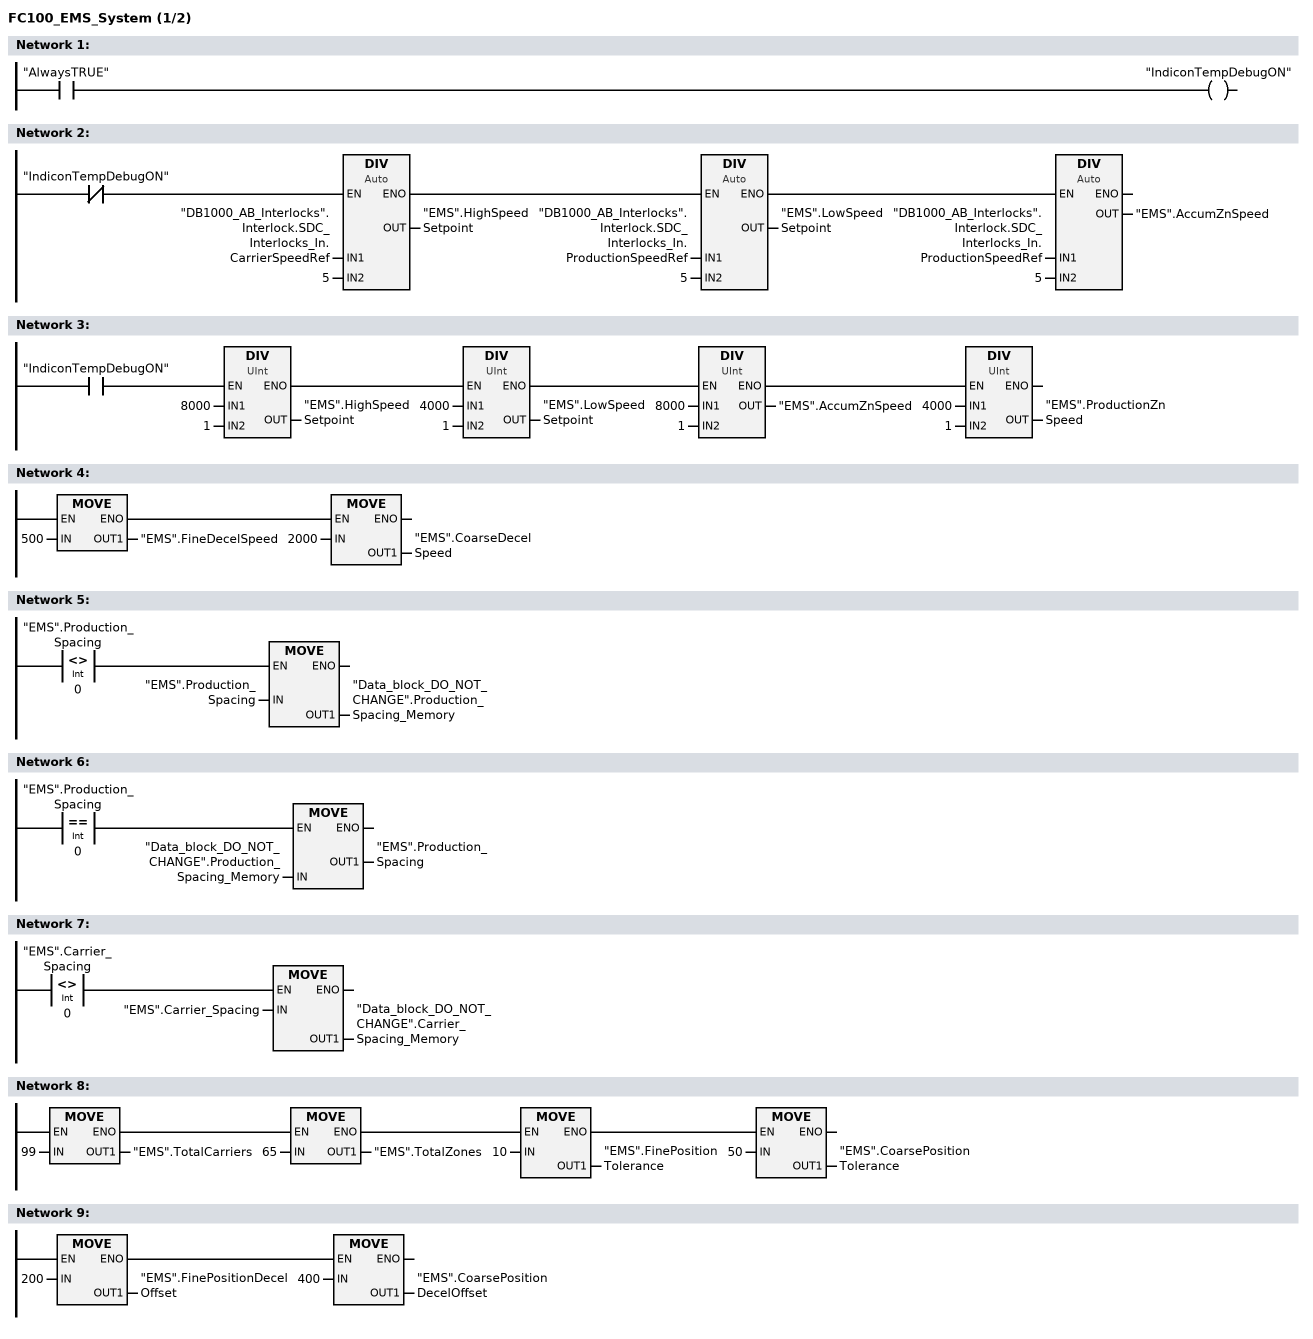
   RUNG wire#powerrail
      Contact( "AlwaysTRUE" )
      Coil( "IndiconTempDebugON" )
   END_RUNG
   // the same network as SCL:
   "IndiconTempDebugON" := "AlwaysTRUE";
END_REGION

REGION Network 2
   RUNG wire#powerrail
      I_Contact( "IndiconTempDebugON" )
      Div(in1 := "DB1000_AB_Interlocks".Interlock.SDC_Interlocks_In.CarrierSpeedRef, in2 := 5, out => "EMS".HighSpeedSetpoint)
      Div(in1 := "DB1000_AB_Interlocks".Interlock.SDC_Interlocks_In.ProductionSpeedRef, in2 := 5, out => "EMS".LowSpeedSetpoint)
      Div(in1 := "DB1000_AB_Interlocks".Interlock.SDC_Interlocks_In.ProductionSpeedRef, in2 := 5, out => "EMS".AccumZnSpeed)
   END_RUNG
   // the same network as SCL:
   IF NOT "IndiconTempDebugON" THEN
       "EMS".HighSpeedSetpoint := "DB1000_AB_Interlocks".Interlock.SDC_Interlocks_In.CarrierSpeedRef / 5;
       "EMS".LowSpeedSetpoint := "DB1000_AB_Interlocks".Interlock.SDC_Interlocks_In.ProductionSpeedRef / 5;
       "EMS".AccumZnSpeed := "DB1000_AB_Interlocks".Interlock.SDC_Interlocks_In.ProductionSpeedRef / 5;
   END_IF;
END_REGION

REGION Network 3
   RUNG wire#powerrail
      Contact( "IndiconTempDebugON" )
      { S7_Templates := "SrcType := UInt" } Div(in1 := 8000, in2 := 1, out => "EMS".HighSpeedSetpoint)
      { S7_Templates := "SrcType := UInt" } Div(in1 := 4000, in2 := 1, out => "EMS".LowSpeedSetpoint)
      { S7_Templates := "SrcType := UInt" } Div(in1 := 8000, in2 := 1, out => "EMS".AccumZnSpeed)
      { S7_Templates := "SrcType := UInt" } Div(in1 := 4000, in2 := 1, out => "EMS".ProductionZnSpeed)
   END_RUNG
   // the same network as SCL:
   IF "IndiconTempDebugON" THEN
       "EMS".HighSpeedSetpoint := 8000 / 1;
       "EMS".LowSpeedSetpoint := 4000 / 1;
       "EMS".AccumZnSpeed := 8000 / 1;
       "EMS".ProductionZnSpeed := 4000 / 1;
   END_IF;
END_REGION

REGION Network 4
   RUNG wire#powerrail
      Move(in := 500, out1 => "EMS".FineDecelSpeed)
      Move(in := 2000, out1 => "EMS".CoarseDecelSpeed)
   END_RUNG
   // the same network as SCL:
   "EMS".FineDecelSpeed := 500;
   "EMS".CoarseDecelSpeed := 2000;
END_REGION

REGION Network 5
   RUNG wire#powerrail
      { S7_Templates := "SrcType := Int" } NE_Contact(in1 := "EMS".Production_Spacing, in2 := 0)
      Move(in := "EMS".Production_Spacing, out1 => "Data_block_DO_NOT_CHANGE".Production_Spacing_Memory)
   END_RUNG
   // the same network as SCL:
   IF "EMS".Production_Spacing <> 0 THEN
       "Data_block_DO_NOT_CHANGE".Production_Spacing_Memory := "EMS".Production_Spacing;
   END_IF;
END_REGION

REGION Network 6
   RUNG wire#powerrail
      { S7_Templates := "SrcType := Int" } EQ_Contact(in1 := "EMS".Production_Spacing, in2 := 0)
      Move(in := "Data_block_DO_NOT_CHANGE".Production_Spacing_Memory, out1 => "EMS".Production_Spacing)
   END_RUNG
   // the same network as SCL:
   IF "EMS".Production_Spacing = 0 THEN
       "EMS".Production_Spacing := "Data_block_DO_NOT_CHANGE".Production_Spacing_Memory;
   END_IF;
END_REGION

REGION Network 7
   RUNG wire#powerrail
      { S7_Templates := "SrcType := Int" } NE_Contact(in1 := "EMS".Carrier_Spacing, in2 := 0)
      Move(in := "EMS".Carrier_Spacing, out1 => "Data_block_DO_NOT_CHANGE".Carrier_Spacing_Memory)
   END_RUNG
   // the same network as SCL:
   IF "EMS".Carrier_Spacing <> 0 THEN
       "Data_block_DO_NOT_CHANGE".Carrier_Spacing_Memory := "EMS".Carrier_Spacing;
   END_IF;
END_REGION

REGION Network 8
   RUNG wire#powerrail
      Move(in := 99, out1 => "EMS".TotalCarriers)
      Move(in := 65, out1 => "EMS".TotalZones)
      Move(in := 10, out1 => "EMS".FinePositionTolerance)
      Move(in := 50, out1 => "EMS".CoarsePositionTolerance)
   END_RUNG
   // the same network as SCL:
   "EMS".TotalCarriers := 99;
   "EMS".TotalZones := 65;
   "EMS".FinePositionTolerance := 10;
   "EMS".CoarsePositionTolerance := 50;
END_REGION

REGION Network 9
   RUNG wire#powerrail
      Move(in := 200, out1 => "EMS".FinePositionDecelOffset)
      Move(in := 400, out1 => "EMS".CoarsePositionDecelOffset)
   END_RUNG
   // the same network as SCL:
   "EMS".FinePositionDecelOffset := 200;
   "EMS".CoarsePositionDecelOffset := 400;
END_REGION

REGION Network 10
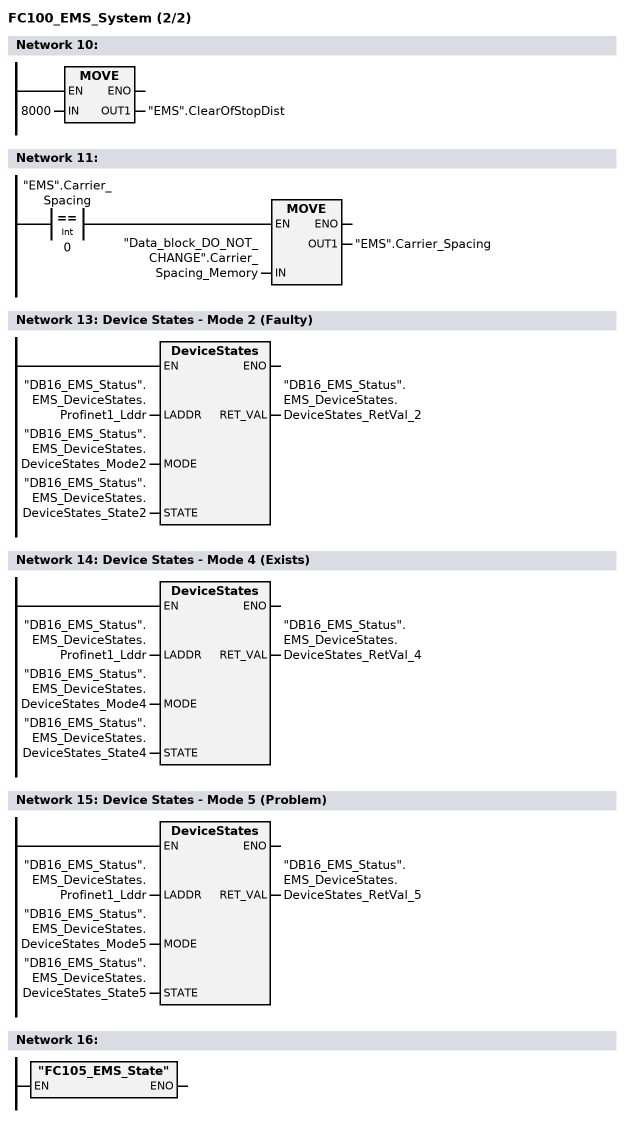
   RUNG wire#powerrail
      Move(in := 8000, out1 => "EMS".ClearOfStopDist)
   END_RUNG
   // the same network as SCL:
   "EMS".ClearOfStopDist := 8000;
END_REGION

REGION Network 11
   RUNG wire#powerrail
      { S7_Templates := "SrcType := Int" } EQ_Contact(in1 := "EMS".Carrier_Spacing, in2 := 0)
      Move(in := "Data_block_DO_NOT_CHANGE".Carrier_Spacing_Memory, out1 => "EMS".Carrier_Spacing)
   END_RUNG
   // the same network as SCL:
   IF "EMS".Carrier_Spacing = 0 THEN
       "EMS".Carrier_Spacing := "Data_block_DO_NOT_CHANGE".Carrier_Spacing_Memory;
   END_IF;
END_REGION

REGION Network 13: Device States - Mode 2 (Faulty)
   // no SCL statement known for DeviceStates: written as a call
   "DB16_EMS_Status".EMS_DeviceStates.DeviceStates_RetVal_2 := DeviceStates(LADDR := "DB16_EMS_Status".EMS_DeviceStates.Profinet1_Lddr,
                           MODE := "DB16_EMS_Status".EMS_DeviceStates.DeviceStates_Mode2,
                           STATE := "DB16_EMS_Status".EMS_DeviceStates.DeviceStates_State2);
END_REGION

REGION Network 14: Device States - Mode 4 (Exists)
   // no SCL statement known for DeviceStates: written as a call
   "DB16_EMS_Status".EMS_DeviceStates.DeviceStates_RetVal_4 := DeviceStates(LADDR := "DB16_EMS_Status".EMS_DeviceStates.Profinet1_Lddr,
                           MODE := "DB16_EMS_Status".EMS_DeviceStates.DeviceStates_Mode4,
                           STATE := "DB16_EMS_Status".EMS_DeviceStates.DeviceStates_State4);
END_REGION

REGION Network 15: Device States - Mode 5 (Problem)
   // no SCL statement known for DeviceStates: written as a call
   "DB16_EMS_Status".EMS_DeviceStates.DeviceStates_RetVal_5 := DeviceStates(LADDR := "DB16_EMS_Status".EMS_DeviceStates.Profinet1_Lddr,
                           MODE := "DB16_EMS_Status".EMS_DeviceStates.DeviceStates_Mode5,
                           STATE := "DB16_EMS_Status".EMS_DeviceStates.DeviceStates_State5);
END_REGION

REGION Network 16
   RUNG wire#powerrail
      "FC105_EMS_State"()
   END_RUNG
   // the same network as SCL:
   "FC105_EMS_State"();
END_REGION
END_FUNCTION

FUNCTION "FC102_TCop_Map_SDCOut" : Void   // FC102, LAD
{ S7_Optimized_Access := 'TRUE' }
VERSION : 0.1
   VAR_TEMP
      tempdisplay : Bool;
      TotalCarriers : Int;
      TotalZones : Int;
      OneShot : Bool;
      countpulse : Bool;
   END_VAR
   VAR_TEMP   // added for the SCL form of the ladder/FBD networks
      _w1 : Bool;
   END_VAR
BEGIN

REGION Network 1
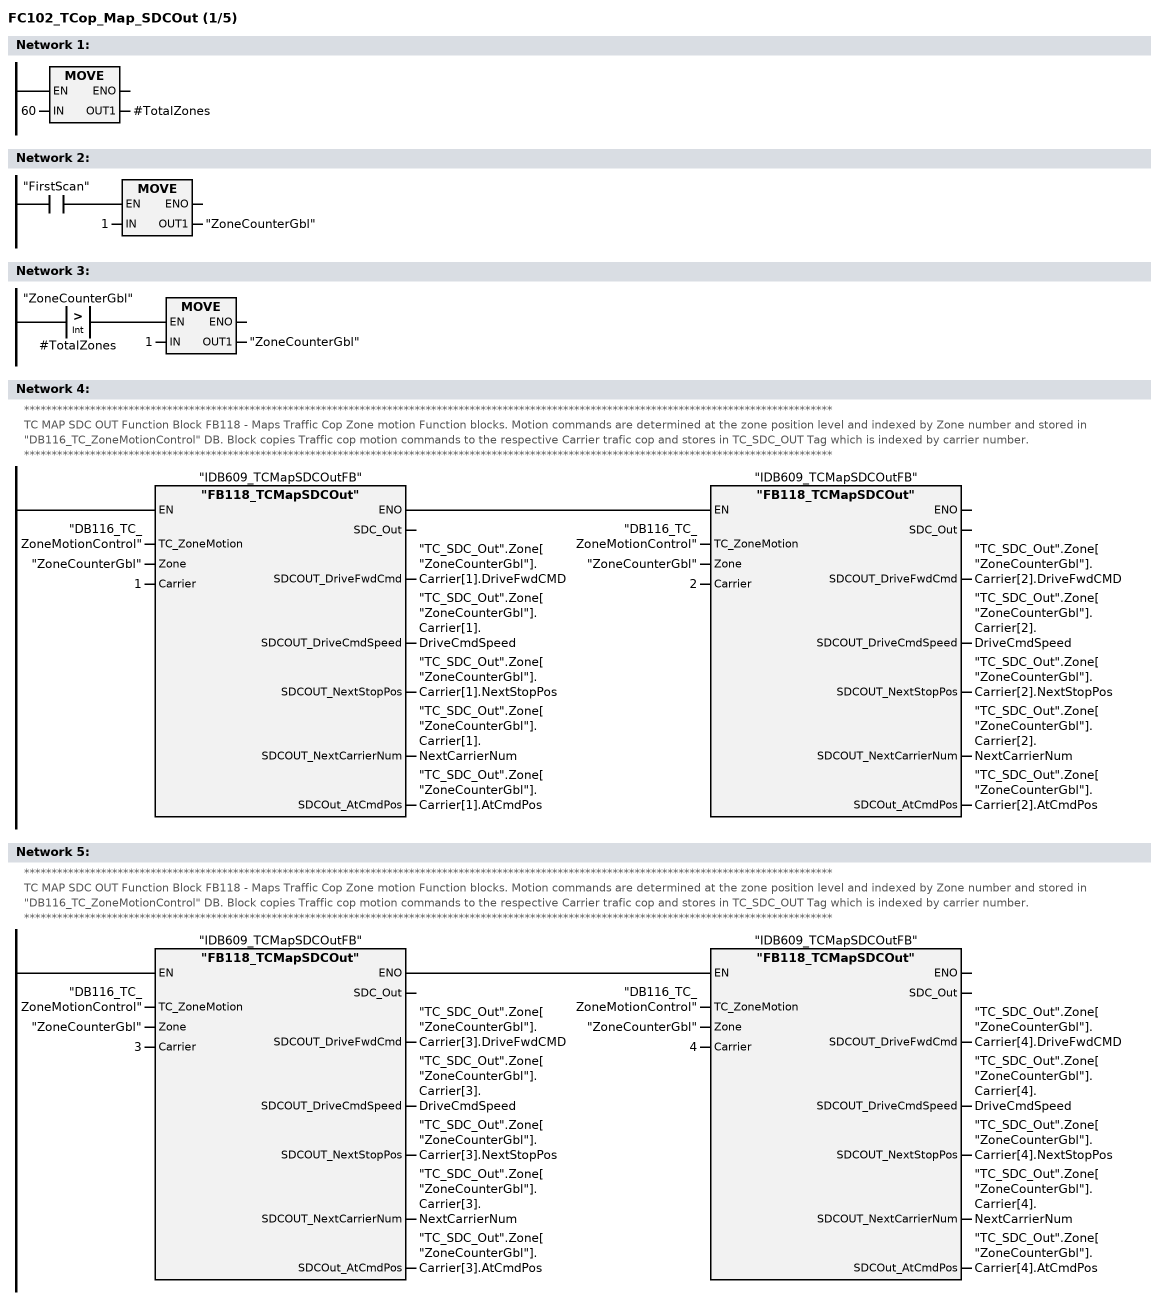
   RUNG wire#powerrail
      Move(in := 60, out1 => #TotalZones)
   END_RUNG
   // the same network as SCL:
   #TotalZones := 60;
END_REGION

REGION Network 2
   RUNG wire#powerrail
      Contact( "FirstScan" )
      Move(in := 1, out1 => "ZoneCounterGbl")
   END_RUNG
   // the same network as SCL:
   IF "FirstScan" THEN "ZoneCounterGbl" := 1; END_IF;
END_REGION

REGION Network 3
   RUNG wire#powerrail
      { S7_Templates := "SrcType := Int" } GT_Contact(in1 := "ZoneCounterGbl", in2 := #TotalZones)
      Move(in := 1, out1 => "ZoneCounterGbl")
   END_RUNG
   // the same network as SCL:
   IF "ZoneCounterGbl" > #TotalZones THEN "ZoneCounterGbl" := 1; END_IF;
END_REGION

REGION Network 4
   // ***************************************************************************************************************************************************
   // 
   // TC MAP SDC OUT Function Block FB118 - Maps Traffic Cop Zone motion Function blocks. Motion commands are determined at the zone position level and indexed by Zone number and stored in 
   //  "DB116_TC_ZoneMotionControl" DB. Block copies Traffic cop motion commands to the respective Carrier trafic cop and stores in TC_SDC_OUT Tag which is indexed by carrier number. 
   // 
   // ***************************************************************************************************************************************************
   RUNG wire#powerrail
      "IDB609_TCMapSDCOutFB"(TC_ZoneMotion := "DB116_TC_ZoneMotionControl", Zone := "ZoneCounterGbl", Carrier := 1, SDC_Out =>, SDCOUT_DriveFwdCmd => "TC_SDC_Out".Zone["ZoneCounterGbl"].Carrier[1].DriveFwdCMD, SDCOUT_DriveCmdSpeed => "TC_SDC_Out".Zone["ZoneCounterGbl"].Carrier[1].DriveCmdSpeed, SDCOUT_NextStopPos => "TC_SDC_Out".Zone["ZoneCounterGbl"].Carrier[1].NextStopPos, SDCOUT_NextCarrierNum => "TC_SDC_Out".Zone["ZoneCounterGbl"].Carrier[1].NextCarrierNum, SDCOut_AtCmdPos => "TC_SDC_Out".Zone["ZoneCounterGbl"].Carrier[1].AtCmdPos)
      "IDB609_TCMapSDCOutFB"(TC_ZoneMotion := "DB116_TC_ZoneMotionControl", Zone := "ZoneCounterGbl", Carrier := 2, SDC_Out =>, SDCOUT_DriveFwdCmd => "TC_SDC_Out".Zone["ZoneCounterGbl"].Carrier[2].DriveFwdCMD, SDCOUT_DriveCmdSpeed => "TC_SDC_Out".Zone["ZoneCounterGbl"].Carrier[2].DriveCmdSpeed, SDCOUT_NextStopPos => "TC_SDC_Out".Zone["ZoneCounterGbl"].Carrier[2].NextStopPos, SDCOUT_NextCarrierNum => "TC_SDC_Out".Zone["ZoneCounterGbl"].Carrier[2].NextCarrierNum, SDCOut_AtCmdPos => "TC_SDC_Out".Zone["ZoneCounterGbl"].Carrier[2].AtCmdPos)
   END_RUNG
   // the same network as SCL:
   "IDB609_TCMapSDCOutFB"(TC_ZoneMotion := "DB116_TC_ZoneMotionControl",   // "FB118_TCMapSDCOut"
                          Zone := "ZoneCounterGbl",
                          Carrier := 1,
                          SDCOUT_DriveFwdCmd => "TC_SDC_Out".Zone["ZoneCounterGbl"].Carrier[1].DriveFwdCMD,
                          SDCOUT_DriveCmdSpeed => "TC_SDC_Out".Zone["ZoneCounterGbl"].Carrier[1].DriveCmdSpeed,
                          SDCOUT_NextStopPos => "TC_SDC_Out".Zone["ZoneCounterGbl"].Carrier[1].NextStopPos,
                          SDCOUT_NextCarrierNum => "TC_SDC_Out".Zone["ZoneCounterGbl"].Carrier[1].NextCarrierNum,
                          SDCOut_AtCmdPos => "TC_SDC_Out".Zone["ZoneCounterGbl"].Carrier[1].AtCmdPos,
                          ENO => #_w1);
   IF #_w1 THEN
       "IDB609_TCMapSDCOutFB"(TC_ZoneMotion := "DB116_TC_ZoneMotionControl",   // "FB118_TCMapSDCOut"
                              Zone := "ZoneCounterGbl",
                              Carrier := 2,
                              SDCOUT_DriveFwdCmd => "TC_SDC_Out".Zone["ZoneCounterGbl"].Carrier[2].DriveFwdCMD,
                              SDCOUT_DriveCmdSpeed => "TC_SDC_Out".Zone["ZoneCounterGbl"].Carrier[2].DriveCmdSpeed,
                              SDCOUT_NextStopPos => "TC_SDC_Out".Zone["ZoneCounterGbl"].Carrier[2].NextStopPos,
                              SDCOUT_NextCarrierNum => "TC_SDC_Out".Zone["ZoneCounterGbl"].Carrier[2].NextCarrierNum,
                              SDCOut_AtCmdPos => "TC_SDC_Out".Zone["ZoneCounterGbl"].Carrier[2].AtCmdPos);
   END_IF;
END_REGION

REGION Network 5
   // ***************************************************************************************************************************************************
   // 
   // TC MAP SDC OUT Function Block FB118 - Maps Traffic Cop Zone motion Function blocks. Motion commands are determined at the zone position level and indexed by Zone number and stored in 
   //  "DB116_TC_ZoneMotionControl" DB. Block copies Traffic cop motion commands to the respective Carrier trafic cop and stores in TC_SDC_OUT Tag which is indexed by carrier number. 
   // 
   // ***************************************************************************************************************************************************
   RUNG wire#powerrail
      "IDB609_TCMapSDCOutFB"(TC_ZoneMotion := "DB116_TC_ZoneMotionControl", Zone := "ZoneCounterGbl", Carrier := 3, SDC_Out =>, SDCOUT_DriveFwdCmd => "TC_SDC_Out".Zone["ZoneCounterGbl"].Carrier[3].DriveFwdCMD, SDCOUT_DriveCmdSpeed => "TC_SDC_Out".Zone["ZoneCounterGbl"].Carrier[3].DriveCmdSpeed, SDCOUT_NextStopPos => "TC_SDC_Out".Zone["ZoneCounterGbl"].Carrier[3].NextStopPos, SDCOUT_NextCarrierNum => "TC_SDC_Out".Zone["ZoneCounterGbl"].Carrier[3].NextCarrierNum, SDCOut_AtCmdPos => "TC_SDC_Out".Zone["ZoneCounterGbl"].Carrier[3].AtCmdPos)
      "IDB609_TCMapSDCOutFB"(TC_ZoneMotion := "DB116_TC_ZoneMotionControl", Zone := "ZoneCounterGbl", Carrier := 4, SDC_Out =>, SDCOUT_DriveFwdCmd => "TC_SDC_Out".Zone["ZoneCounterGbl"].Carrier[4].DriveFwdCMD, SDCOUT_DriveCmdSpeed => "TC_SDC_Out".Zone["ZoneCounterGbl"].Carrier[4].DriveCmdSpeed, SDCOUT_NextStopPos => "TC_SDC_Out".Zone["ZoneCounterGbl"].Carrier[4].NextStopPos, SDCOUT_NextCarrierNum => "TC_SDC_Out".Zone["ZoneCounterGbl"].Carrier[4].NextCarrierNum, SDCOut_AtCmdPos => "TC_SDC_Out".Zone["ZoneCounterGbl"].Carrier[4].AtCmdPos)
   END_RUNG
   // the same network as SCL:
   "IDB609_TCMapSDCOutFB"(TC_ZoneMotion := "DB116_TC_ZoneMotionControl",   // "FB118_TCMapSDCOut"
                          Zone := "ZoneCounterGbl",
                          Carrier := 3,
                          SDCOUT_DriveFwdCmd => "TC_SDC_Out".Zone["ZoneCounterGbl"].Carrier[3].DriveFwdCMD,
                          SDCOUT_DriveCmdSpeed => "TC_SDC_Out".Zone["ZoneCounterGbl"].Carrier[3].DriveCmdSpeed,
                          SDCOUT_NextStopPos => "TC_SDC_Out".Zone["ZoneCounterGbl"].Carrier[3].NextStopPos,
                          SDCOUT_NextCarrierNum => "TC_SDC_Out".Zone["ZoneCounterGbl"].Carrier[3].NextCarrierNum,
                          SDCOut_AtCmdPos => "TC_SDC_Out".Zone["ZoneCounterGbl"].Carrier[3].AtCmdPos,
                          ENO => #_w1);
   IF #_w1 THEN
       "IDB609_TCMapSDCOutFB"(TC_ZoneMotion := "DB116_TC_ZoneMotionControl",   // "FB118_TCMapSDCOut"
                              Zone := "ZoneCounterGbl",
                              Carrier := 4,
                              SDCOUT_DriveFwdCmd => "TC_SDC_Out".Zone["ZoneCounterGbl"].Carrier[4].DriveFwdCMD,
                              SDCOUT_DriveCmdSpeed => "TC_SDC_Out".Zone["ZoneCounterGbl"].Carrier[4].DriveCmdSpeed,
                              SDCOUT_NextStopPos => "TC_SDC_Out".Zone["ZoneCounterGbl"].Carrier[4].NextStopPos,
                              SDCOUT_NextCarrierNum => "TC_SDC_Out".Zone["ZoneCounterGbl"].Carrier[4].NextCarrierNum,
                              SDCOut_AtCmdPos => "TC_SDC_Out".Zone["ZoneCounterGbl"].Carrier[4].AtCmdPos);
   END_IF;
END_REGION

REGION Network 6
   // ***************************************************************************************************************************************************
   // 
   // TC MAP SDC OUT Function Block FB118 - Maps Traffic Cop Zone motion Function blocks. Motion commands are determined at the zone position level and indexed by Zone number and stored in 
   //  "DB116_TC_ZoneMotionControl" DB. Block copies Traffic cop motion commands to the respective Carrier trafic cop and stores in TC_SDC_OUT Tag which is indexed by carrier number. 
   // 
   // ***************************************************************************************************************************************************
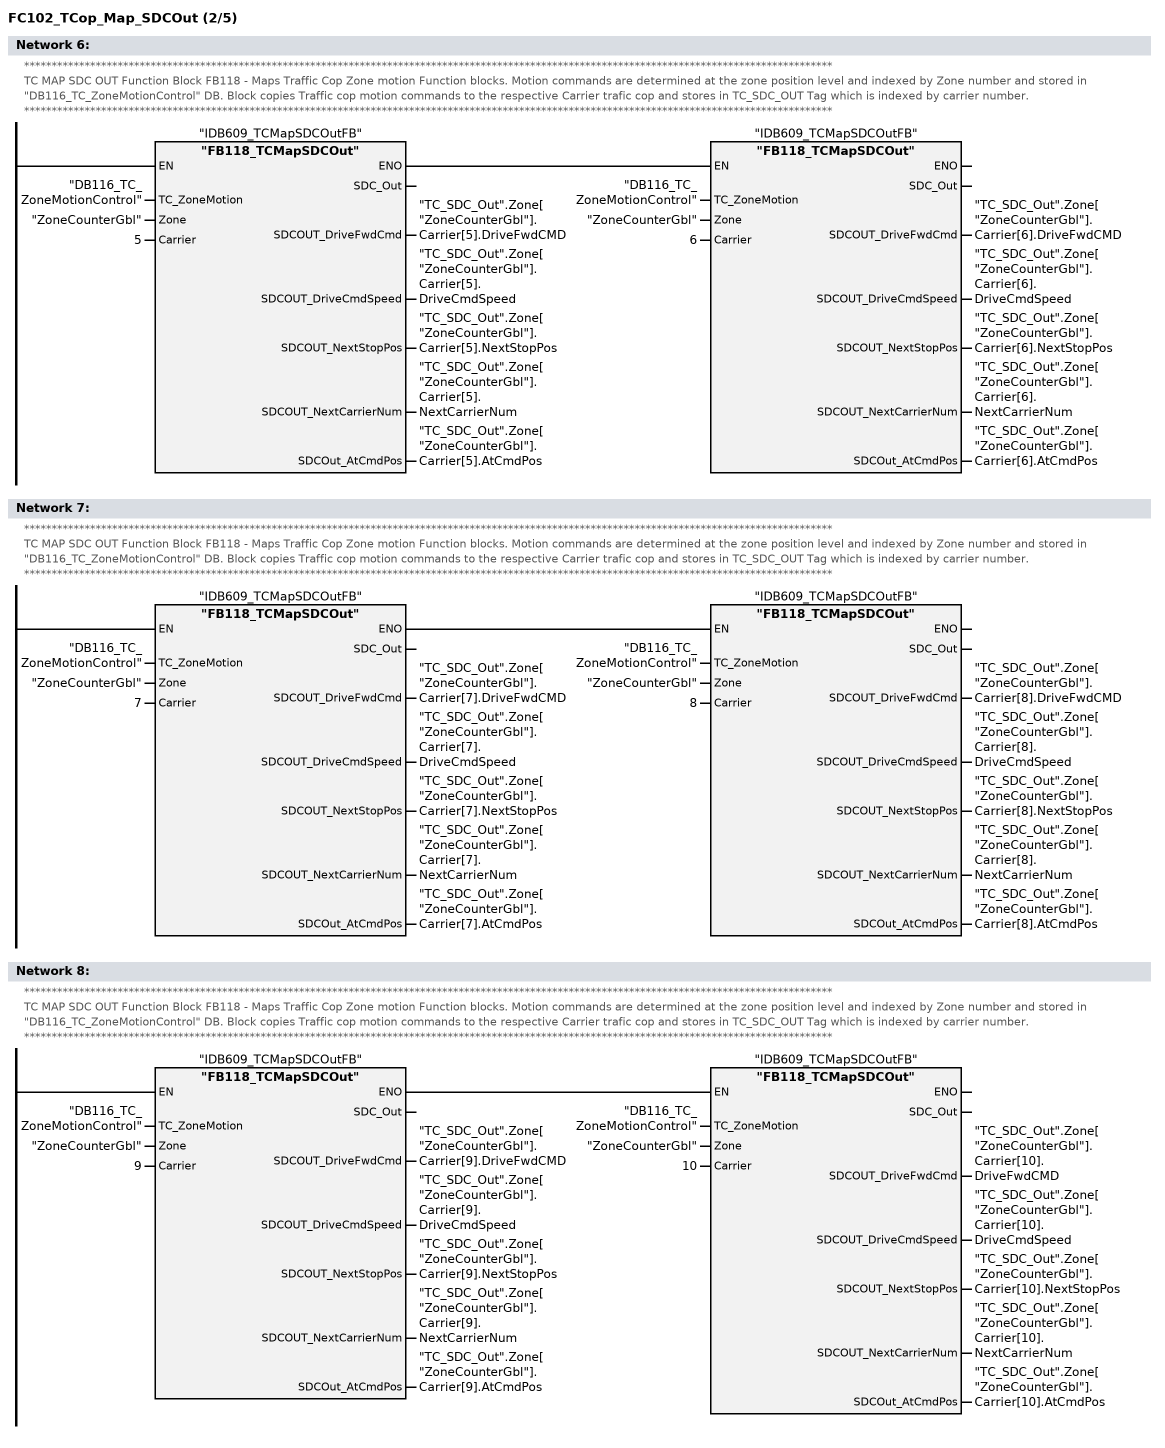
   RUNG wire#powerrail
      "IDB609_TCMapSDCOutFB"(TC_ZoneMotion := "DB116_TC_ZoneMotionControl", Zone := "ZoneCounterGbl", Carrier := 5, SDC_Out =>, SDCOUT_DriveFwdCmd => "TC_SDC_Out".Zone["ZoneCounterGbl"].Carrier[5].DriveFwdCMD, SDCOUT_DriveCmdSpeed => "TC_SDC_Out".Zone["ZoneCounterGbl"].Carrier[5].DriveCmdSpeed, SDCOUT_NextStopPos => "TC_SDC_Out".Zone["ZoneCounterGbl"].Carrier[5].NextStopPos, SDCOUT_NextCarrierNum => "TC_SDC_Out".Zone["ZoneCounterGbl"].Carrier[5].NextCarrierNum, SDCOut_AtCmdPos => "TC_SDC_Out".Zone["ZoneCounterGbl"].Carrier[5].AtCmdPos)
      "IDB609_TCMapSDCOutFB"(TC_ZoneMotion := "DB116_TC_ZoneMotionControl", Zone := "ZoneCounterGbl", Carrier := 6, SDC_Out =>, SDCOUT_DriveFwdCmd => "TC_SDC_Out".Zone["ZoneCounterGbl"].Carrier[6].DriveFwdCMD, SDCOUT_DriveCmdSpeed => "TC_SDC_Out".Zone["ZoneCounterGbl"].Carrier[6].DriveCmdSpeed, SDCOUT_NextStopPos => "TC_SDC_Out".Zone["ZoneCounterGbl"].Carrier[6].NextStopPos, SDCOUT_NextCarrierNum => "TC_SDC_Out".Zone["ZoneCounterGbl"].Carrier[6].NextCarrierNum, SDCOut_AtCmdPos => "TC_SDC_Out".Zone["ZoneCounterGbl"].Carrier[6].AtCmdPos)
   END_RUNG
   // the same network as SCL:
   "IDB609_TCMapSDCOutFB"(TC_ZoneMotion := "DB116_TC_ZoneMotionControl",   // "FB118_TCMapSDCOut"
                          Zone := "ZoneCounterGbl",
                          Carrier := 5,
                          SDCOUT_DriveFwdCmd => "TC_SDC_Out".Zone["ZoneCounterGbl"].Carrier[5].DriveFwdCMD,
                          SDCOUT_DriveCmdSpeed => "TC_SDC_Out".Zone["ZoneCounterGbl"].Carrier[5].DriveCmdSpeed,
                          SDCOUT_NextStopPos => "TC_SDC_Out".Zone["ZoneCounterGbl"].Carrier[5].NextStopPos,
                          SDCOUT_NextCarrierNum => "TC_SDC_Out".Zone["ZoneCounterGbl"].Carrier[5].NextCarrierNum,
                          SDCOut_AtCmdPos => "TC_SDC_Out".Zone["ZoneCounterGbl"].Carrier[5].AtCmdPos,
                          ENO => #_w1);
   IF #_w1 THEN
       "IDB609_TCMapSDCOutFB"(TC_ZoneMotion := "DB116_TC_ZoneMotionControl",   // "FB118_TCMapSDCOut"
                              Zone := "ZoneCounterGbl",
                              Carrier := 6,
                              SDCOUT_DriveFwdCmd => "TC_SDC_Out".Zone["ZoneCounterGbl"].Carrier[6].DriveFwdCMD,
                              SDCOUT_DriveCmdSpeed => "TC_SDC_Out".Zone["ZoneCounterGbl"].Carrier[6].DriveCmdSpeed,
                              SDCOUT_NextStopPos => "TC_SDC_Out".Zone["ZoneCounterGbl"].Carrier[6].NextStopPos,
                              SDCOUT_NextCarrierNum => "TC_SDC_Out".Zone["ZoneCounterGbl"].Carrier[6].NextCarrierNum,
                              SDCOut_AtCmdPos => "TC_SDC_Out".Zone["ZoneCounterGbl"].Carrier[6].AtCmdPos);
   END_IF;
END_REGION

REGION Network 7
   // ***************************************************************************************************************************************************
   // 
   // TC MAP SDC OUT Function Block FB118 - Maps Traffic Cop Zone motion Function blocks. Motion commands are determined at the zone position level and indexed by Zone number and stored in 
   //  "DB116_TC_ZoneMotionControl" DB. Block copies Traffic cop motion commands to the respective Carrier trafic cop and stores in TC_SDC_OUT Tag which is indexed by carrier number. 
   // 
   // ***************************************************************************************************************************************************
   RUNG wire#powerrail
      "IDB609_TCMapSDCOutFB"(TC_ZoneMotion := "DB116_TC_ZoneMotionControl", Zone := "ZoneCounterGbl", Carrier := 7, SDC_Out =>, SDCOUT_DriveFwdCmd => "TC_SDC_Out".Zone["ZoneCounterGbl"].Carrier[7].DriveFwdCMD, SDCOUT_DriveCmdSpeed => "TC_SDC_Out".Zone["ZoneCounterGbl"].Carrier[7].DriveCmdSpeed, SDCOUT_NextStopPos => "TC_SDC_Out".Zone["ZoneCounterGbl"].Carrier[7].NextStopPos, SDCOUT_NextCarrierNum => "TC_SDC_Out".Zone["ZoneCounterGbl"].Carrier[7].NextCarrierNum, SDCOut_AtCmdPos => "TC_SDC_Out".Zone["ZoneCounterGbl"].Carrier[7].AtCmdPos)
      "IDB609_TCMapSDCOutFB"(TC_ZoneMotion := "DB116_TC_ZoneMotionControl", Zone := "ZoneCounterGbl", Carrier := 8, SDC_Out =>, SDCOUT_DriveFwdCmd => "TC_SDC_Out".Zone["ZoneCounterGbl"].Carrier[8].DriveFwdCMD, SDCOUT_DriveCmdSpeed => "TC_SDC_Out".Zone["ZoneCounterGbl"].Carrier[8].DriveCmdSpeed, SDCOUT_NextStopPos => "TC_SDC_Out".Zone["ZoneCounterGbl"].Carrier[8].NextStopPos, SDCOUT_NextCarrierNum => "TC_SDC_Out".Zone["ZoneCounterGbl"].Carrier[8].NextCarrierNum, SDCOut_AtCmdPos => "TC_SDC_Out".Zone["ZoneCounterGbl"].Carrier[8].AtCmdPos)
   END_RUNG
   // the same network as SCL:
   "IDB609_TCMapSDCOutFB"(TC_ZoneMotion := "DB116_TC_ZoneMotionControl",   // "FB118_TCMapSDCOut"
                          Zone := "ZoneCounterGbl",
                          Carrier := 7,
                          SDCOUT_DriveFwdCmd => "TC_SDC_Out".Zone["ZoneCounterGbl"].Carrier[7].DriveFwdCMD,
                          SDCOUT_DriveCmdSpeed => "TC_SDC_Out".Zone["ZoneCounterGbl"].Carrier[7].DriveCmdSpeed,
                          SDCOUT_NextStopPos => "TC_SDC_Out".Zone["ZoneCounterGbl"].Carrier[7].NextStopPos,
                          SDCOUT_NextCarrierNum => "TC_SDC_Out".Zone["ZoneCounterGbl"].Carrier[7].NextCarrierNum,
                          SDCOut_AtCmdPos => "TC_SDC_Out".Zone["ZoneCounterGbl"].Carrier[7].AtCmdPos,
                          ENO => #_w1);
   IF #_w1 THEN
       "IDB609_TCMapSDCOutFB"(TC_ZoneMotion := "DB116_TC_ZoneMotionControl",   // "FB118_TCMapSDCOut"
                              Zone := "ZoneCounterGbl",
                              Carrier := 8,
                              SDCOUT_DriveFwdCmd => "TC_SDC_Out".Zone["ZoneCounterGbl"].Carrier[8].DriveFwdCMD,
                              SDCOUT_DriveCmdSpeed => "TC_SDC_Out".Zone["ZoneCounterGbl"].Carrier[8].DriveCmdSpeed,
                              SDCOUT_NextStopPos => "TC_SDC_Out".Zone["ZoneCounterGbl"].Carrier[8].NextStopPos,
                              SDCOUT_NextCarrierNum => "TC_SDC_Out".Zone["ZoneCounterGbl"].Carrier[8].NextCarrierNum,
                              SDCOut_AtCmdPos => "TC_SDC_Out".Zone["ZoneCounterGbl"].Carrier[8].AtCmdPos);
   END_IF;
END_REGION

REGION Network 8
   // ***************************************************************************************************************************************************
   // 
   // TC MAP SDC OUT Function Block FB118 - Maps Traffic Cop Zone motion Function blocks. Motion commands are determined at the zone position level and indexed by Zone number and stored in 
   //  "DB116_TC_ZoneMotionControl" DB. Block copies Traffic cop motion commands to the respective Carrier trafic cop and stores in TC_SDC_OUT Tag which is indexed by carrier number. 
   // 
   // ***************************************************************************************************************************************************
   RUNG wire#powerrail
      "IDB609_TCMapSDCOutFB"(TC_ZoneMotion := "DB116_TC_ZoneMotionControl", Zone := "ZoneCounterGbl", Carrier := 9, SDC_Out =>, SDCOUT_DriveFwdCmd => "TC_SDC_Out".Zone["ZoneCounterGbl"].Carrier[9].DriveFwdCMD, SDCOUT_DriveCmdSpeed => "TC_SDC_Out".Zone["ZoneCounterGbl"].Carrier[9].DriveCmdSpeed, SDCOUT_NextStopPos => "TC_SDC_Out".Zone["ZoneCounterGbl"].Carrier[9].NextStopPos, SDCOUT_NextCarrierNum => "TC_SDC_Out".Zone["ZoneCounterGbl"].Carrier[9].NextCarrierNum, SDCOut_AtCmdPos => "TC_SDC_Out".Zone["ZoneCounterGbl"].Carrier[9].AtCmdPos)
      "IDB609_TCMapSDCOutFB"(TC_ZoneMotion := "DB116_TC_ZoneMotionControl", Zone := "ZoneCounterGbl", Carrier := 10, SDC_Out =>, SDCOUT_DriveFwdCmd => "TC_SDC_Out".Zone["ZoneCounterGbl"].Carrier[10].DriveFwdCMD, SDCOUT_DriveCmdSpeed => "TC_SDC_Out".Zone["ZoneCounterGbl"].Carrier[10].DriveCmdSpeed, SDCOUT_NextStopPos => "TC_SDC_Out".Zone["ZoneCounterGbl"].Carrier[10].NextStopPos, SDCOUT_NextCarrierNum => "TC_SDC_Out".Zone["ZoneCounterGbl"].Carrier[10].NextCarrierNum, SDCOut_AtCmdPos => "TC_SDC_Out".Zone["ZoneCounterGbl"].Carrier[10].AtCmdPos)
   END_RUNG
   // the same network as SCL:
   "IDB609_TCMapSDCOutFB"(TC_ZoneMotion := "DB116_TC_ZoneMotionControl",   // "FB118_TCMapSDCOut"
                          Zone := "ZoneCounterGbl",
                          Carrier := 9,
                          SDCOUT_DriveFwdCmd => "TC_SDC_Out".Zone["ZoneCounterGbl"].Carrier[9].DriveFwdCMD,
                          SDCOUT_DriveCmdSpeed => "TC_SDC_Out".Zone["ZoneCounterGbl"].Carrier[9].DriveCmdSpeed,
                          SDCOUT_NextStopPos => "TC_SDC_Out".Zone["ZoneCounterGbl"].Carrier[9].NextStopPos,
                          SDCOUT_NextCarrierNum => "TC_SDC_Out".Zone["ZoneCounterGbl"].Carrier[9].NextCarrierNum,
                          SDCOut_AtCmdPos => "TC_SDC_Out".Zone["ZoneCounterGbl"].Carrier[9].AtCmdPos,
                          ENO => #_w1);
   IF #_w1 THEN
       "IDB609_TCMapSDCOutFB"(TC_ZoneMotion := "DB116_TC_ZoneMotionControl",   // "FB118_TCMapSDCOut"
                              Zone := "ZoneCounterGbl",
                              Carrier := 10,
                              SDCOUT_DriveFwdCmd => "TC_SDC_Out".Zone["ZoneCounterGbl"].Carrier[10].DriveFwdCMD,
                              SDCOUT_DriveCmdSpeed => "TC_SDC_Out".Zone["ZoneCounterGbl"].Carrier[10].DriveCmdSpeed,
                              SDCOUT_NextStopPos => "TC_SDC_Out".Zone["ZoneCounterGbl"].Carrier[10].NextStopPos,
                              SDCOUT_NextCarrierNum => "TC_SDC_Out".Zone["ZoneCounterGbl"].Carrier[10].NextCarrierNum,
                              SDCOut_AtCmdPos => "TC_SDC_Out".Zone["ZoneCounterGbl"].Carrier[10].AtCmdPos);
   END_IF;
END_REGION

REGION Network 9
   // ***************************************************************************************************************************************************
   // 
   // TC MAP SDC OUT Function Block FB118 - Maps Traffic Cop Zone motion Function blocks. Motion commands are determined at the zone position level and indexed by Zone number and stored in 
   //  "DB116_TC_ZoneMotionControl" DB. Block copies Traffic cop motion commands to the respective Carrier trafic cop and stores in TC_SDC_OUT Tag which is indexed by carrier number. 
   // 
   // ***************************************************************************************************************************************************
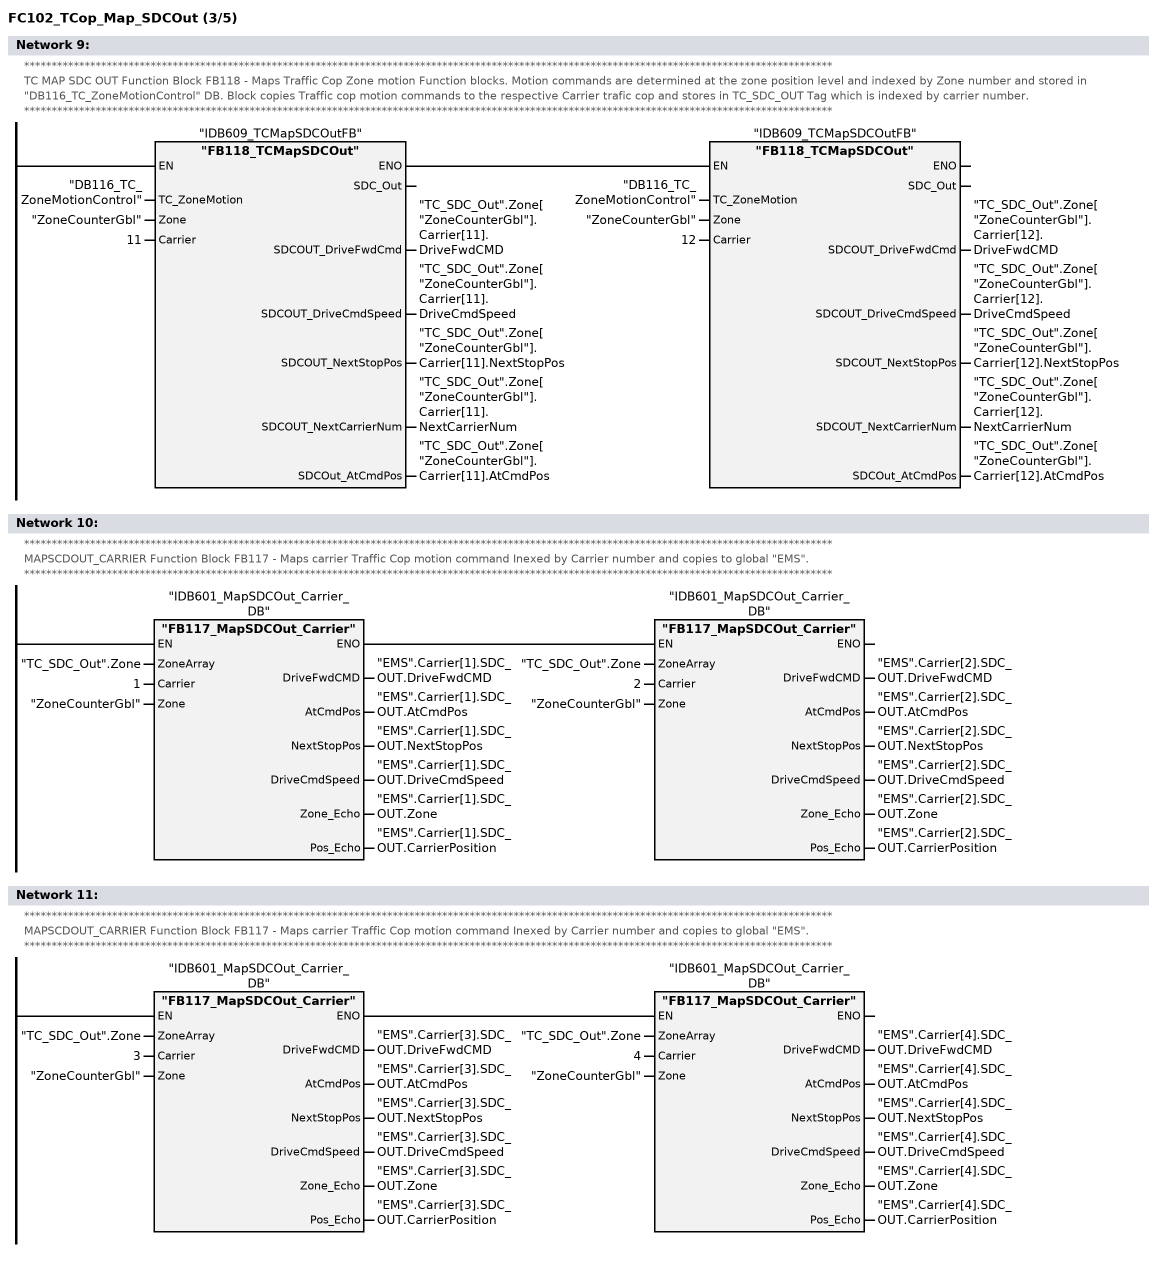
   RUNG wire#powerrail
      "IDB609_TCMapSDCOutFB"(TC_ZoneMotion := "DB116_TC_ZoneMotionControl", Zone := "ZoneCounterGbl", Carrier := 11, SDC_Out =>, SDCOUT_DriveFwdCmd => "TC_SDC_Out".Zone["ZoneCounterGbl"].Carrier[11].DriveFwdCMD, SDCOUT_DriveCmdSpeed => "TC_SDC_Out".Zone["ZoneCounterGbl"].Carrier[11].DriveCmdSpeed, SDCOUT_NextStopPos => "TC_SDC_Out".Zone["ZoneCounterGbl"].Carrier[11].NextStopPos, SDCOUT_NextCarrierNum => "TC_SDC_Out".Zone["ZoneCounterGbl"].Carrier[11].NextCarrierNum, SDCOut_AtCmdPos => "TC_SDC_Out".Zone["ZoneCounterGbl"].Carrier[11].AtCmdPos)
      "IDB609_TCMapSDCOutFB"(TC_ZoneMotion := "DB116_TC_ZoneMotionControl", Zone := "ZoneCounterGbl", Carrier := 12, SDC_Out =>, SDCOUT_DriveFwdCmd => "TC_SDC_Out".Zone["ZoneCounterGbl"].Carrier[12].DriveFwdCMD, SDCOUT_DriveCmdSpeed => "TC_SDC_Out".Zone["ZoneCounterGbl"].Carrier[12].DriveCmdSpeed, SDCOUT_NextStopPos => "TC_SDC_Out".Zone["ZoneCounterGbl"].Carrier[12].NextStopPos, SDCOUT_NextCarrierNum => "TC_SDC_Out".Zone["ZoneCounterGbl"].Carrier[12].NextCarrierNum, SDCOut_AtCmdPos => "TC_SDC_Out".Zone["ZoneCounterGbl"].Carrier[12].AtCmdPos)
   END_RUNG
   // the same network as SCL:
   "IDB609_TCMapSDCOutFB"(TC_ZoneMotion := "DB116_TC_ZoneMotionControl",   // "FB118_TCMapSDCOut"
                          Zone := "ZoneCounterGbl",
                          Carrier := 11,
                          SDCOUT_DriveFwdCmd => "TC_SDC_Out".Zone["ZoneCounterGbl"].Carrier[11].DriveFwdCMD,
                          SDCOUT_DriveCmdSpeed => "TC_SDC_Out".Zone["ZoneCounterGbl"].Carrier[11].DriveCmdSpeed,
                          SDCOUT_NextStopPos => "TC_SDC_Out".Zone["ZoneCounterGbl"].Carrier[11].NextStopPos,
                          SDCOUT_NextCarrierNum => "TC_SDC_Out".Zone["ZoneCounterGbl"].Carrier[11].NextCarrierNum,
                          SDCOut_AtCmdPos => "TC_SDC_Out".Zone["ZoneCounterGbl"].Carrier[11].AtCmdPos,
                          ENO => #_w1);
   IF #_w1 THEN
       "IDB609_TCMapSDCOutFB"(TC_ZoneMotion := "DB116_TC_ZoneMotionControl",   // "FB118_TCMapSDCOut"
                              Zone := "ZoneCounterGbl",
                              Carrier := 12,
                              SDCOUT_DriveFwdCmd => "TC_SDC_Out".Zone["ZoneCounterGbl"].Carrier[12].DriveFwdCMD,
                              SDCOUT_DriveCmdSpeed => "TC_SDC_Out".Zone["ZoneCounterGbl"].Carrier[12].DriveCmdSpeed,
                              SDCOUT_NextStopPos => "TC_SDC_Out".Zone["ZoneCounterGbl"].Carrier[12].NextStopPos,
                              SDCOUT_NextCarrierNum => "TC_SDC_Out".Zone["ZoneCounterGbl"].Carrier[12].NextCarrierNum,
                              SDCOut_AtCmdPos => "TC_SDC_Out".Zone["ZoneCounterGbl"].Carrier[12].AtCmdPos);
   END_IF;
END_REGION

REGION Network 10
   // ***************************************************************************************************************************************************
   // 
   // MAPSCDOUT_CARRIER Function Block FB117 - Maps carrier Traffic Cop motion command Inexed by Carrier number and copies to global "EMS". 
   // 
   // ***************************************************************************************************************************************************
   RUNG wire#powerrail
      "IDB601_MapSDCOut_Carrier_DB"(ZoneArray := "TC_SDC_Out".Zone, Carrier := 1, Zone := "ZoneCounterGbl", DriveFwdCMD => "EMS".Carrier[1].SDC_OUT.DriveFwdCMD, AtCmdPos => "EMS".Carrier[1].SDC_OUT.AtCmdPos, NextStopPos => "EMS".Carrier[1].SDC_OUT.NextStopPos, DriveCmdSpeed => "EMS".Carrier[1].SDC_OUT.DriveCmdSpeed, Zone_Echo => "EMS".Carrier[1].SDC_OUT.Zone, Pos_Echo => "EMS".Carrier[1].SDC_OUT.CarrierPosition)
      "IDB601_MapSDCOut_Carrier_DB"(ZoneArray := "TC_SDC_Out".Zone, Carrier := 2, Zone := "ZoneCounterGbl", DriveFwdCMD => "EMS".Carrier[2].SDC_OUT.DriveFwdCMD, AtCmdPos => "EMS".Carrier[2].SDC_OUT.AtCmdPos, NextStopPos => "EMS".Carrier[2].SDC_OUT.NextStopPos, DriveCmdSpeed => "EMS".Carrier[2].SDC_OUT.DriveCmdSpeed, Zone_Echo => "EMS".Carrier[2].SDC_OUT.Zone, Pos_Echo => "EMS".Carrier[2].SDC_OUT.CarrierPosition)
   END_RUNG
   // the same network as SCL:
   "IDB601_MapSDCOut_Carrier_DB"(ZoneArray := "TC_SDC_Out".Zone,   // "FB117_MapSDCOut_Carrier"
                           Carrier := 1,
                           Zone := "ZoneCounterGbl",
                           DriveFwdCMD => "EMS".Carrier[1].SDC_OUT.DriveFwdCMD,
                           AtCmdPos => "EMS".Carrier[1].SDC_OUT.AtCmdPos,
                           NextStopPos => "EMS".Carrier[1].SDC_OUT.NextStopPos,
                           DriveCmdSpeed => "EMS".Carrier[1].SDC_OUT.DriveCmdSpeed,
                           Zone_Echo => "EMS".Carrier[1].SDC_OUT.Zone,
                           Pos_Echo => "EMS".Carrier[1].SDC_OUT.CarrierPosition,
                           ENO => #_w1);
   IF #_w1 THEN
       "IDB601_MapSDCOut_Carrier_DB"(ZoneArray := "TC_SDC_Out".Zone,   // "FB117_MapSDCOut_Carrier"
                               Carrier := 2,
                               Zone := "ZoneCounterGbl",
                               DriveFwdCMD => "EMS".Carrier[2].SDC_OUT.DriveFwdCMD,
                               AtCmdPos => "EMS".Carrier[2].SDC_OUT.AtCmdPos,
                               NextStopPos => "EMS".Carrier[2].SDC_OUT.NextStopPos,
                               DriveCmdSpeed => "EMS".Carrier[2].SDC_OUT.DriveCmdSpeed,
                               Zone_Echo => "EMS".Carrier[2].SDC_OUT.Zone,
                               Pos_Echo => "EMS".Carrier[2].SDC_OUT.CarrierPosition);
   END_IF;
END_REGION

REGION Network 11
   // ***************************************************************************************************************************************************
   // 
   // MAPSCDOUT_CARRIER Function Block FB117 - Maps carrier Traffic Cop motion command Inexed by Carrier number and copies to global "EMS". 
   // 
   // ***************************************************************************************************************************************************
   RUNG wire#powerrail
      "IDB601_MapSDCOut_Carrier_DB"(ZoneArray := "TC_SDC_Out".Zone, Carrier := 3, Zone := "ZoneCounterGbl", DriveFwdCMD => "EMS".Carrier[3].SDC_OUT.DriveFwdCMD, AtCmdPos => "EMS".Carrier[3].SDC_OUT.AtCmdPos, NextStopPos => "EMS".Carrier[3].SDC_OUT.NextStopPos, DriveCmdSpeed => "EMS".Carrier[3].SDC_OUT.DriveCmdSpeed, Zone_Echo => "EMS".Carrier[3].SDC_OUT.Zone, Pos_Echo => "EMS".Carrier[3].SDC_OUT.CarrierPosition)
      "IDB601_MapSDCOut_Carrier_DB"(ZoneArray := "TC_SDC_Out".Zone, Carrier := 4, Zone := "ZoneCounterGbl", DriveFwdCMD => "EMS".Carrier[4].SDC_OUT.DriveFwdCMD, AtCmdPos => "EMS".Carrier[4].SDC_OUT.AtCmdPos, NextStopPos => "EMS".Carrier[4].SDC_OUT.NextStopPos, DriveCmdSpeed => "EMS".Carrier[4].SDC_OUT.DriveCmdSpeed, Zone_Echo => "EMS".Carrier[4].SDC_OUT.Zone, Pos_Echo => "EMS".Carrier[4].SDC_OUT.CarrierPosition)
   END_RUNG
   // the same network as SCL:
   "IDB601_MapSDCOut_Carrier_DB"(ZoneArray := "TC_SDC_Out".Zone,   // "FB117_MapSDCOut_Carrier"
                           Carrier := 3,
                           Zone := "ZoneCounterGbl",
                           DriveFwdCMD => "EMS".Carrier[3].SDC_OUT.DriveFwdCMD,
                           AtCmdPos => "EMS".Carrier[3].SDC_OUT.AtCmdPos,
                           NextStopPos => "EMS".Carrier[3].SDC_OUT.NextStopPos,
                           DriveCmdSpeed => "EMS".Carrier[3].SDC_OUT.DriveCmdSpeed,
                           Zone_Echo => "EMS".Carrier[3].SDC_OUT.Zone,
                           Pos_Echo => "EMS".Carrier[3].SDC_OUT.CarrierPosition,
                           ENO => #_w1);
   IF #_w1 THEN
       "IDB601_MapSDCOut_Carrier_DB"(ZoneArray := "TC_SDC_Out".Zone,   // "FB117_MapSDCOut_Carrier"
                               Carrier := 4,
                               Zone := "ZoneCounterGbl",
                               DriveFwdCMD => "EMS".Carrier[4].SDC_OUT.DriveFwdCMD,
                               AtCmdPos => "EMS".Carrier[4].SDC_OUT.AtCmdPos,
                               NextStopPos => "EMS".Carrier[4].SDC_OUT.NextStopPos,
                               DriveCmdSpeed => "EMS".Carrier[4].SDC_OUT.DriveCmdSpeed,
                               Zone_Echo => "EMS".Carrier[4].SDC_OUT.Zone,
                               Pos_Echo => "EMS".Carrier[4].SDC_OUT.CarrierPosition);
   END_IF;
END_REGION

REGION Network 12
   // ***************************************************************************************************************************************************
   // 
   // MAPSCDOUT_CARRIER Function Block FB117 - Maps carrier Traffic Cop motion command Inexed by Carrier number and copies to global "EMS". 
   // 
   // ***************************************************************************************************************************************************
